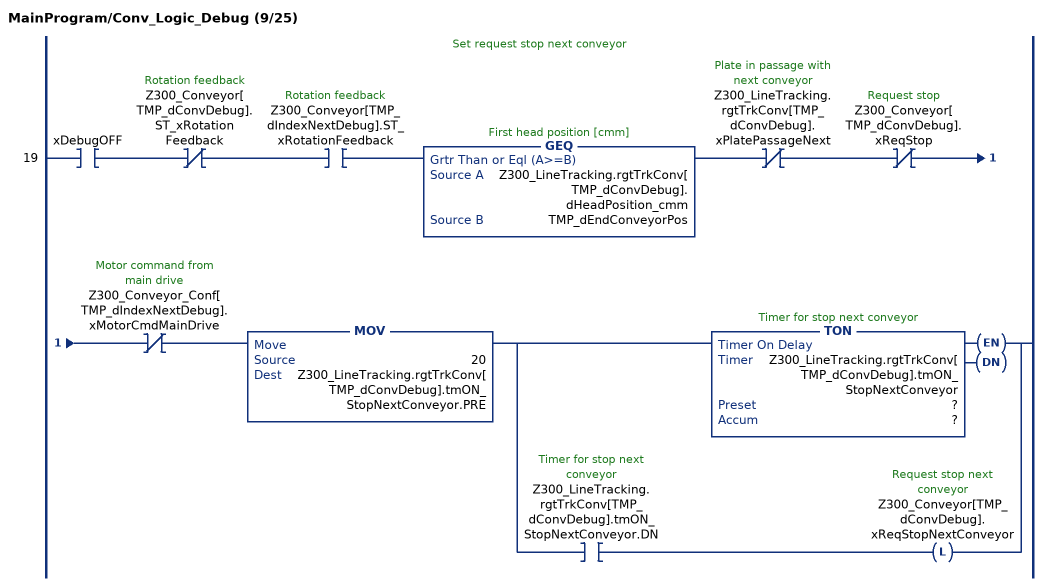
   // Set request stop next conveyor
   19: XIC(xDebugOFF)XIO(Z300_Conveyor[TMP_dConvDebug].ST_xRotationFeedback)XIC(Z300_Conveyor[TMP_dIndexNextDebug].ST_xRotationFeedback)GEQ(Z300_LineTracking.rgtTrkConv[TMP_dConvDebug].dHeadPosition_cmm,TMP_dEndConveyorPos)XIO(Z300_LineTracking.rgtTrkConv[TMP_dConvDebug].xPlatePassageNext)XIO(Z300_Conveyor[TMP_dConvDebug].xReqStop)XIO(Z300_Conveyor_Conf[TMP_dIndexNextDebug].xMotorCmdMainDrive)MOV(20,Z300_LineTracking.rgtTrkConv[TMP_dConvDebug].tmON_StopNextConveyor.PRE)[TON(Z300_LineTracking.rgtTrkConv[TMP_dConvDebug].tmON_StopNextConveyor,?,?) ,XIC(Z300_LineTracking.rgtTrkConv[TMP_dConvDebug].tmON_StopNextConveyor.DN) OTL(Z300_Conveyor[TMP_dConvDebug].xReqStopNextConveyor) ];
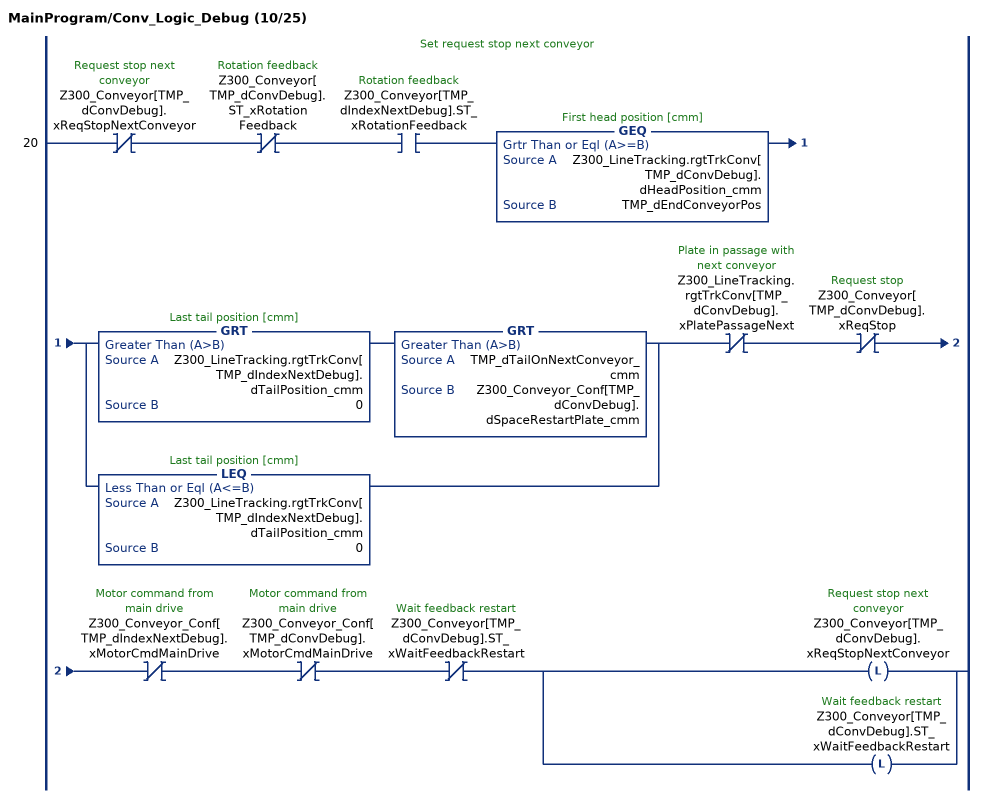
   // Set request stop next conveyor
   20: XIO(Z300_Conveyor[TMP_dConvDebug].xReqStopNextConveyor)XIO(Z300_Conveyor[TMP_dConvDebug].ST_xRotationFeedback)XIC(Z300_Conveyor[TMP_dIndexNextDebug].ST_xRotationFeedback)GEQ(Z300_LineTracking.rgtTrkConv[TMP_dConvDebug].dHeadPosition_cmm,TMP_dEndConveyorPos)[GRT(Z300_LineTracking.rgtTrkConv[TMP_dIndexNextDebug].dTailPosition_cmm,0) GRT(TMP_dTailOnNextConveyor_cmm,Z300_Conveyor_Conf[TMP_dConvDebug].dSpaceRestartPlate_cmm) ,LEQ(Z300_LineTracking.rgtTrkConv[TMP_dIndexNextDebug].dTailPosition_cmm,0) ]XIO(Z300_LineTracking.rgtTrkConv[TMP_dConvDebug].xPlatePassageNext)XIO(Z300_Conveyor[TMP_dConvDebug].xReqStop)XIO(Z300_Conveyor_Conf[TMP_dIndexNextDebug].xMotorCmdMainDrive)XIO(Z300_Conveyor_Conf[TMP_dConvDebug].xMotorCmdMainDrive)XIO(Z300_Conveyor[TMP_dConvDebug].ST_xWaitFeedbackRestart)[OTL(Z300_Conveyor[TMP_dConvDebug].xReqStopNextConveyor) ,OTL(Z300_Conveyor[TMP_dConvDebug].ST_xWaitFeedbackRestart) ];
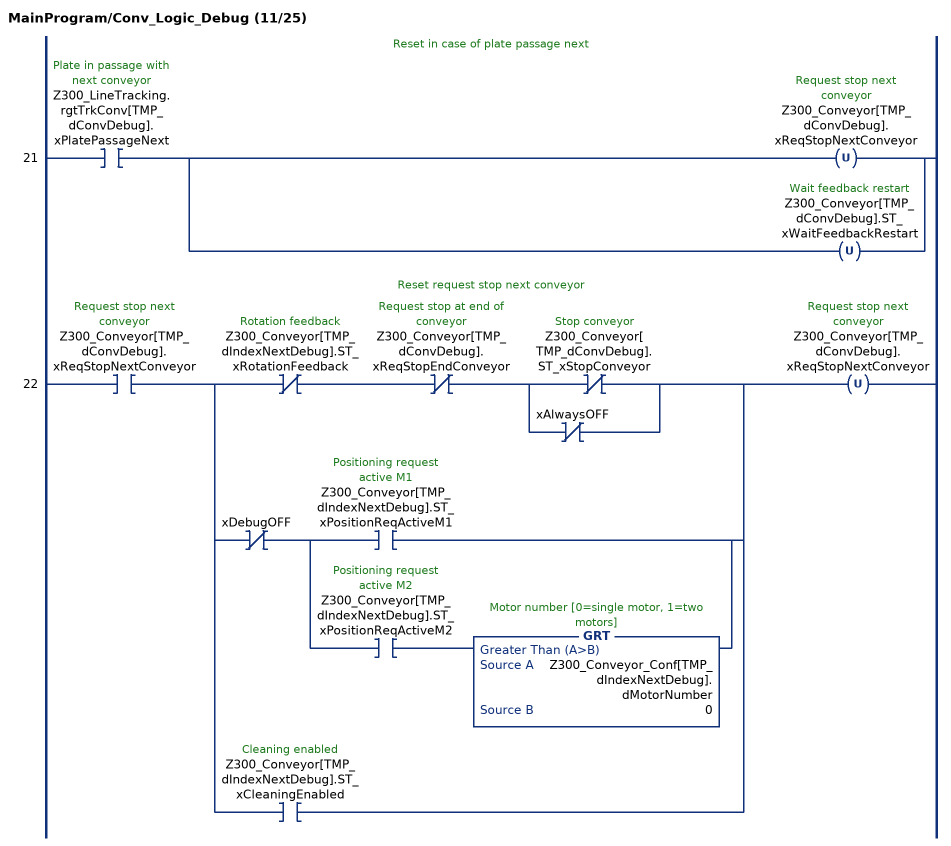
   // Reset in case of plate passage next
   21: XIC(Z300_LineTracking.rgtTrkConv[TMP_dConvDebug].xPlatePassageNext)[OTU(Z300_Conveyor[TMP_dConvDebug].xReqStopNextConveyor) ,OTU(Z300_Conveyor[TMP_dConvDebug].ST_xWaitFeedbackRestart) ];
   // Reset request stop next conveyor
   22: XIC(Z300_Conveyor[TMP_dConvDebug].xReqStopNextConveyor)[XIO(Z300_Conveyor[TMP_dIndexNextDebug].ST_xRotationFeedback) XIO(Z300_Conveyor[TMP_dConvDebug].xReqStopEndConveyor) [XIO(Z300_Conveyor[TMP_dConvDebug].ST_xStopConveyor) ,XIO(xAlwaysOFF) ] ,XIO(xDebugOFF) [XIC(Z300_Conveyor[TMP_dIndexNextDebug].ST_xPositionReqActiveM1) ,XIC(Z300_Conveyor[TMP_dIndexNextDebug].ST_xPositionReqActiveM2) GRT(Z300_Conveyor_Conf[TMP_dIndexNextDebug].dMotorNumber,0) ] ,XIC(Z300_Conveyor[TMP_dIndexNextDebug].ST_xCleaningEnabled) ]OTU(Z300_Conveyor[TMP_dConvDebug].xReqStopNextConveyor);
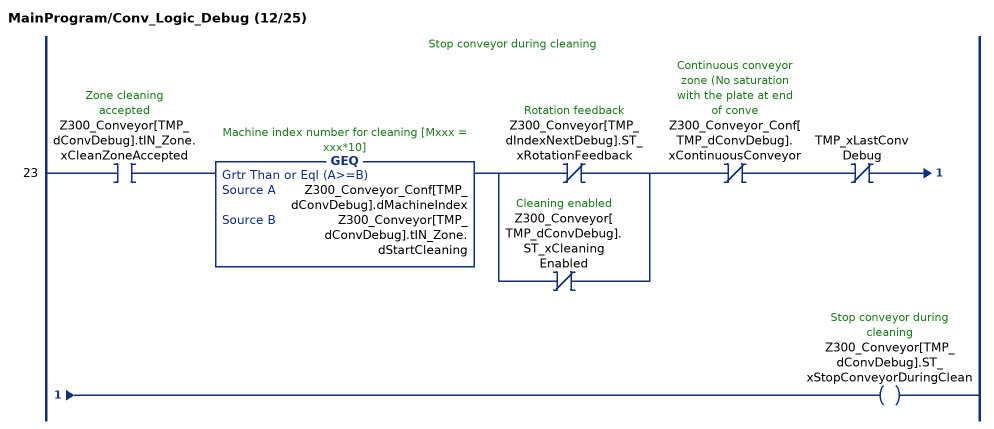
   // Stop conveyor during cleaning
   23: XIC(Z300_Conveyor[TMP_dConvDebug].tIN_Zone.xCleanZoneAccepted)GEQ(Z300_Conveyor_Conf[TMP_dConvDebug].dMachineIndex,Z300_Conveyor[TMP_dConvDebug].tIN_Zone.dStartCleaning)[XIO(Z300_Conveyor[TMP_dIndexNextDebug].ST_xRotationFeedback) ,XIO(Z300_Conveyor[TMP_dConvDebug].ST_xCleaningEnabled) ]XIO(Z300_Conveyor_Conf[TMP_dConvDebug].xContinuousConveyor)XIO(TMP_xLastConvDebug)OTE(Z300_Conveyor[TMP_dConvDebug].ST_xStopConveyorDuringClean);
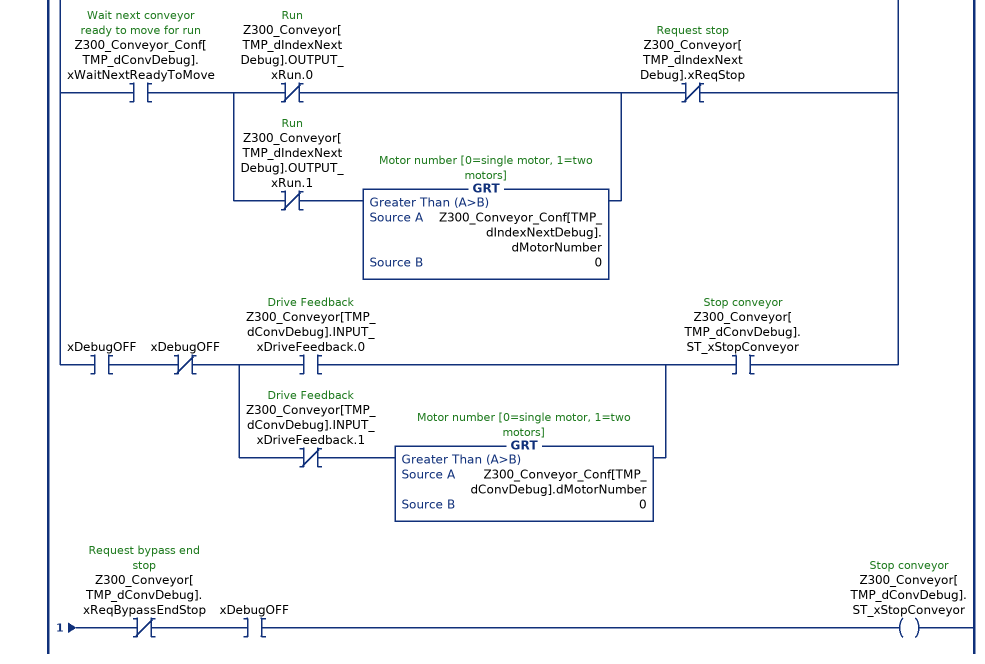
   // Stop conveyor
   24: [[XIC(Z300_LineTracking.rgtTrkConv[TMP_dConvDebug].xPlatePassagePrevious) [XIO(Z300_Conveyor[TMP_dIndexPreviousDebug].ST_xOutputEnable) ,XIC(Z300_Conveyor[TMP_dIndexPreviousDebug].ST_xWaitStopConveyor) ,XIC(xAlwaysOFF) XIC(Z300_Conveyor[TMP_dIndexPreviousDebug].xReqStop) ] ,XIC(Z300_LineTracking.rgtTrkConv[TMP_dConvDebug].xPlatePassageNext) XIO(TMP_xLastConvDebug) [XIO(Z300_Conveyor[TMP_dIndexNextDebug].ST_xOutMotorRun) ,XIO(Z300_Conveyor[TMP_dIndexNextDebug].INPUT_xSafetyConveyor) ] ,XIC(Z300_Conveyor[TMP_dConvDebug].ST_xStopPlateAtEndConveyor) ,XIC(Z300_Conveyor[TMP_dConvDebug].xReqStopNextConveyor) XIC(Z300_Conveyor[TMP_dIndexNextDebug].ST_xRotationFeedback) ,XIC(Z300_Conveyor[TMP_dConvDebug].ST_xStopConveyorDuringClean) ] [XIO(Z300_Conveyor_Conf[TMP_dConvDebug].xContinuousConveyor) ,XIC(Z300_Conveyor_Conf[TMP_dConvDebug].xEnableStopPlateContinuousZone) XIC(Z300_Conveyor[TMP_dConvDebug].xReqStopEndConveyor) ] ,XIC(Z300_Conveyor[TMP_dIndexPreviousDebug].xReqStopNextConveyor) XIO(Z300_Conveyor[TMP_dConvDebug].tIN_Zone.xCleanZoneAccepted) XIO(Z300_LineTracking.rgtTrkConv[TMP_dConvDebug].xGlassPresence) ,XIC(Z300_Conveyor_Conf[TMP_dConvDebug].xWaitNextReadyToMove) [XIO(Z300_Conveyor[TMP_dIndexNextDebug].OUTPUT_xRun.0) ,XIO(Z300_Conveyor[TMP_dIndexNextDebug].OUTPUT_xRun.1) GRT(Z300_Conveyor_Conf[TMP_dIndexNextDebug].dMotorNumber,0) ] XIO(Z300_Conveyor[TMP_dIndexNextDebug].xReqStop) ,XIC(xDebugOFF) XIO(xDebugOFF) [XIC(Z300_Conveyor[TMP_dConvDebug].INPUT_xDriveFeedback.0) ,XIO(Z300_Conveyor[TMP_dConvDebug].INPUT_xDriveFeedback.1) GRT(Z300_Conveyor_Conf[TMP_dConvDebug].dMotorNumber,0) ] XIC(Z300_Conveyor[TMP_dConvDebug].ST_xStopConveyor) ]XIO(Z300_Conveyor[TMP_dConvDebug].xReqBypassEndStop)XIC(xDebugOFF)OTE(Z300_Conveyor[TMP_dConvDebug].ST_xStopConveyor);
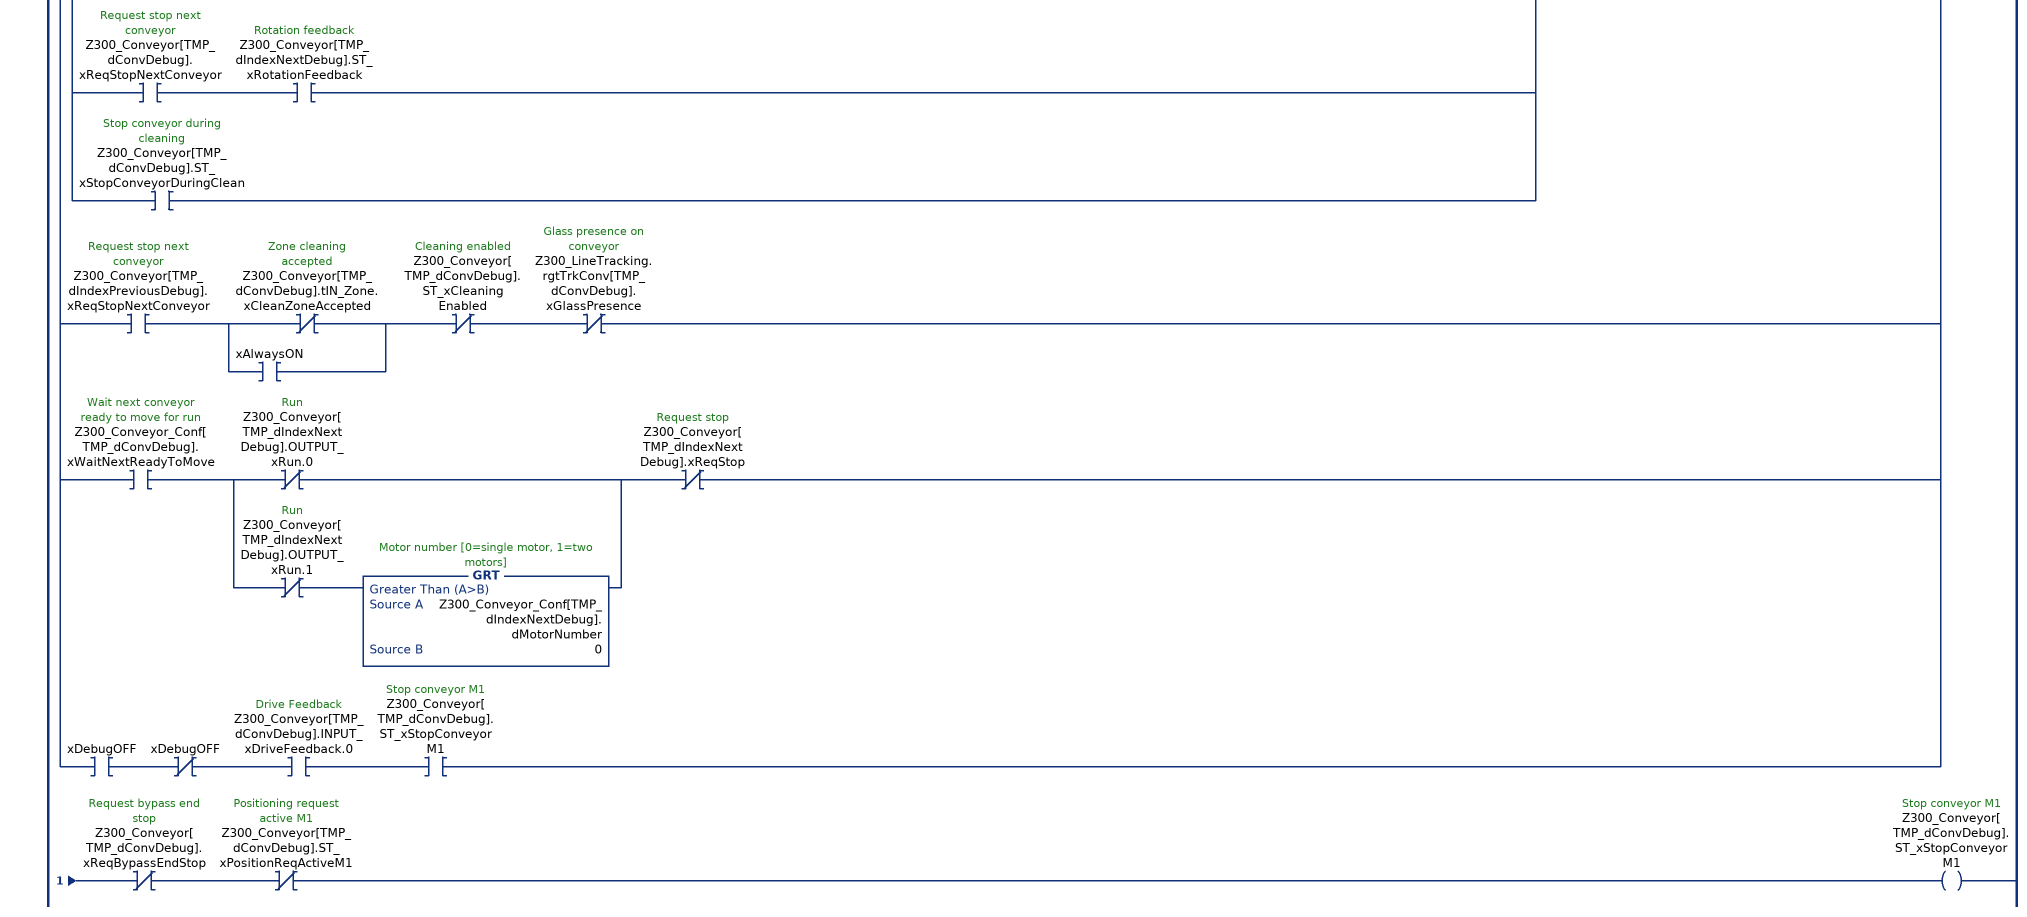
   // Stop conveyor M1
   // Monterrey VF2 - If this is conveyor after drop section I stop convveyor just if tail is under certain quote
   25: [[XIC(Z300_LineTracking.rgtTrkConv[TMP_dConvDebug].xPlatePassagePrevious) [XIO(Z300_Conveyor[TMP_dIndexPreviousDebug].ST_xOutputEnable) ,XIC(xDebugOFF) XIO(Z300_Conveyor[TMP_dIndexPreviousDebug].tmON_DelayReadyToMove[0].DN) ,XIC(Z300_Conveyor[TMP_dIndexPreviousDebug].ST_xInitialCondition) ,XIC(xDebugOFF) XIC(Z300_Conveyor[TMP_dIndexPreviousDebug].ST_xWaitStopConveyor) ,XIC(xAlwaysOFF) XIC(Z300_Conveyor[TMP_dIndexPreviousDebug].xReqStop) ] ,XIC(Z300_LineTracking.rgtTrkConv[TMP_dConvDebug].xPlatePassageNext) XIO(TMP_xLastConvDebug) [XIO(xDebugOFF) [EQU(TMP_dConvDebug,12) LES(Z300_LineTracking.rgtTrkConv[TMP_dConvDebug].dTailPosition_cmm,4100000) ,NEQ(TMP_dConvDebug,12) ] XIO(xDebugOFF) [XIO(Z300_Conveyor[TMP_dIndexNextDebug].ST_xOutMotorRun) ,XIC(xAlwaysON) ] XIO(Z300_Conveyor[TMP_dIndexNextDebug].ST_rgxConveyorOutRunSgm.0) XIO(Z300_Conveyor[TMP_dIndexNextDebug].ST_rgxConveyorOutRunSgm.1) ,XIO(Z300_Conveyor[TMP_dIndexNextDebug].INPUT_xSafetyConveyor) ] ,XIC(Z300_Conveyor[TMP_dConvDebug].ST_xStopPlateAtEndConveyor) XIO(Z300_Conveyor[TMP_dConvDebug].xReqBypassEndConveyorM1) ,XIC(Z300_Conveyor[TMP_dConvDebug].xReqStopNextConveyor) XIC(Z300_Conveyor[TMP_dIndexNextDebug].ST_xRotationFeedback) ,XIC(Z300_Conveyor[TMP_dConvDebug].ST_xStopConveyorDuringClean) ] [XIO(Z300_Conveyor_Conf[TMP_dConvDebug].xContinuousConveyor) ,XIC(Z300_Conveyor_Conf[TMP_dConvDebug].xEnableStopPlateContinuousZone) XIC(Z300_Conveyor[TMP_dConvDebug].xReqStopEndConveyor) ] ,XIC(Z300_Conveyor[TMP_dIndexPreviousDebug].xReqStopNextConveyor) [XIO(Z300_Conveyor[TMP_dConvDebug].tIN_Zone.xCleanZoneAccepted) ,XIC(xAlwaysON) ] XIO(Z300_Conveyor[TMP_dConvDebug].ST_xCleaningEnabled) XIO(Z300_LineTracking.rgtTrkConv[TMP_dConvDebug].xGlassPresence) ,XIC(Z300_Conveyor_Conf[TMP_dConvDebug].xWaitNextReadyToMove) [XIO(Z300_Conveyor[TMP_dIndexNextDebug].OUTPUT_xRun.0) ,XIO(Z300_Conveyor[TMP_dIndexNextDebug].OUTPUT_xRun.1) GRT(Z300_Conveyor_Conf[TMP_dIndexNextDebug].dMotorNumber,0) ] XIO(Z300_Conveyor[TMP_dIndexNextDebug].xReqStop) ,XIC(xDebugOFF) XIO(xDebugOFF) XIC(Z300_Conveyor[TMP_dConvDebug].INPUT_xDriveFeedback.0) XIC(Z300_Conveyor[TMP_dConvDebug].ST_xStopConveyorM1) ]XIO(Z300_Conveyor[TMP_dConvDebug].xReqBypassEndStop)XIO(Z300_Conveyor[TMP_dConvDebug].ST_xPositionReqActiveM1)OTE(Z300_Conveyor[TMP_dConvDebug].ST_xStopConveyorM1);
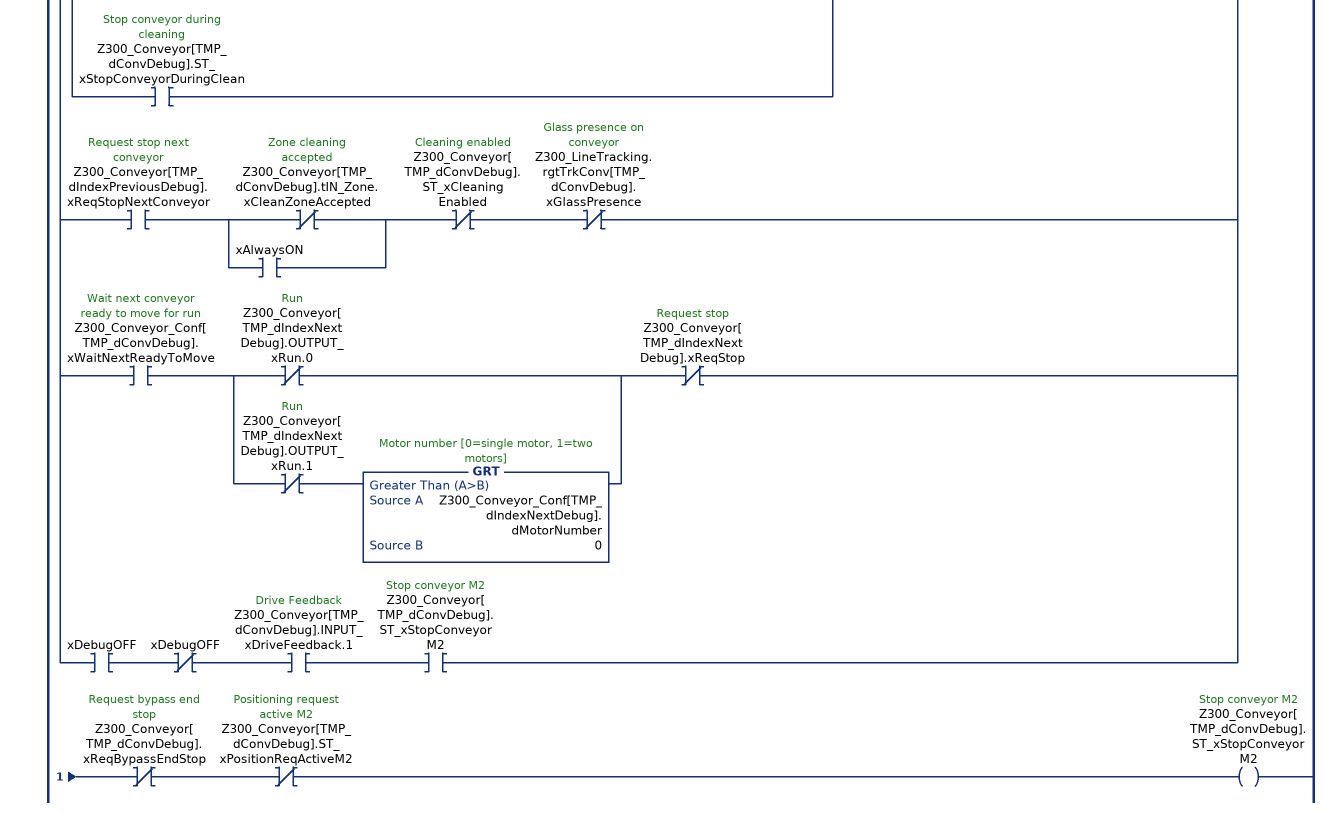
   // Stop conveyor M2
   // Monterrey VF2 - If this is conveyor after drop section I stop convveyor just if tail is under certain quote
   26: [[XIC(Z300_LineTracking.rgtTrkConv[TMP_dConvDebug].xPlatePassagePrevious) [XIO(Z300_Conveyor[TMP_dIndexPreviousDebug].ST_xOutputEnable) ,XIC(xDebugOFF) XIO(Z300_Conveyor[TMP_dIndexPreviousDebug].tmON_DelayReadyToMove[1].DN) ,XIC(Z300_Conveyor[TMP_dIndexPreviousDebug].ST_xInitialCondition) ,XIC(xDebugOFF) XIC(Z300_Conveyor[TMP_dIndexPreviousDebug].ST_xWaitStopConveyor) ,XIC(xAlwaysOFF) XIC(Z300_Conveyor[TMP_dIndexPreviousDebug].xReqStop) ] ,XIC(Z300_LineTracking.rgtTrkConv[TMP_dConvDebug].xPlatePassageNext) XIO(TMP_xLastConvDebug) [[XIO(Z300_Conveyor[TMP_dIndexNextDebug].ST_xOutMotorRun) ,XIC(xAlwaysON) ] XIO(Z300_Conveyor[TMP_dIndexNextDebug].ST_rgxConveyorOutRunSgm.0) XIO(Z300_Conveyor[TMP_dIndexNextDebug].ST_rgxConveyorOutRunSgm.1) ,XIO(Z300_Conveyor[TMP_dIndexNextDebug].INPUT_xSafetyConveyor) ] ,XIC(Z300_Conveyor[TMP_dConvDebug].ST_xStopPlateAtEndConveyor) XIO(Z300_Conveyor[TMP_dConvDebug].xReqBypassEndConveyorM2) ,XIC(Z300_Conveyor[TMP_dConvDebug].xReqStopNextConveyor) XIC(Z300_Conveyor[TMP_dIndexNextDebug].ST_xRotationFeedback) ,XIC(Z300_Conveyor[TMP_dConvDebug].ST_xStopConveyorDuringClean) ] [XIO(Z300_Conveyor_Conf[TMP_dConvDebug].xContinuousConveyor) ,XIC(Z300_Conveyor_Conf[TMP_dConvDebug].xEnableStopPlateContinuousZone) XIC(Z300_Conveyor[TMP_dConvDebug].xReqStopEndConveyor) ] ,XIC(Z300_Conveyor[TMP_dIndexPreviousDebug].xReqStopNextConveyor) [XIO(Z300_Conveyor[TMP_dConvDebug].tIN_Zone.xCleanZoneAccepted) ,XIC(xAlwaysON) ] XIO(Z300_Conveyor[TMP_dConvDebug].ST_xCleaningEnabled) XIO(Z300_LineTracking.rgtTrkConv[TMP_dConvDebug].xGlassPresence) ,XIC(Z300_Conveyor_Conf[TMP_dConvDebug].xWaitNextReadyToMove) [XIO(Z300_Conveyor[TMP_dIndexNextDebug].OUTPUT_xRun.0) ,XIO(Z300_Conveyor[TMP_dIndexNextDebug].OUTPUT_xRun.1) GRT(Z300_Conveyor_Conf[TMP_dIndexNextDebug].dMotorNumber,0) ] XIO(Z300_Conveyor[TMP_dIndexNextDebug].xReqStop) ,XIC(xDebugOFF) XIO(xDebugOFF) XIC(Z300_Conveyor[TMP_dConvDebug].INPUT_xDriveFeedback.1) XIC(Z300_Conveyor[TMP_dConvDebug].ST_xStopConveyorM2) ]XIO(Z300_Conveyor[TMP_dConvDebug].xReqBypassEndStop)XIO(Z300_Conveyor[TMP_dConvDebug].ST_xPositionReqActiveM2)OTE(Z300_Conveyor[TMP_dConvDebug].ST_xStopConveyorM2);
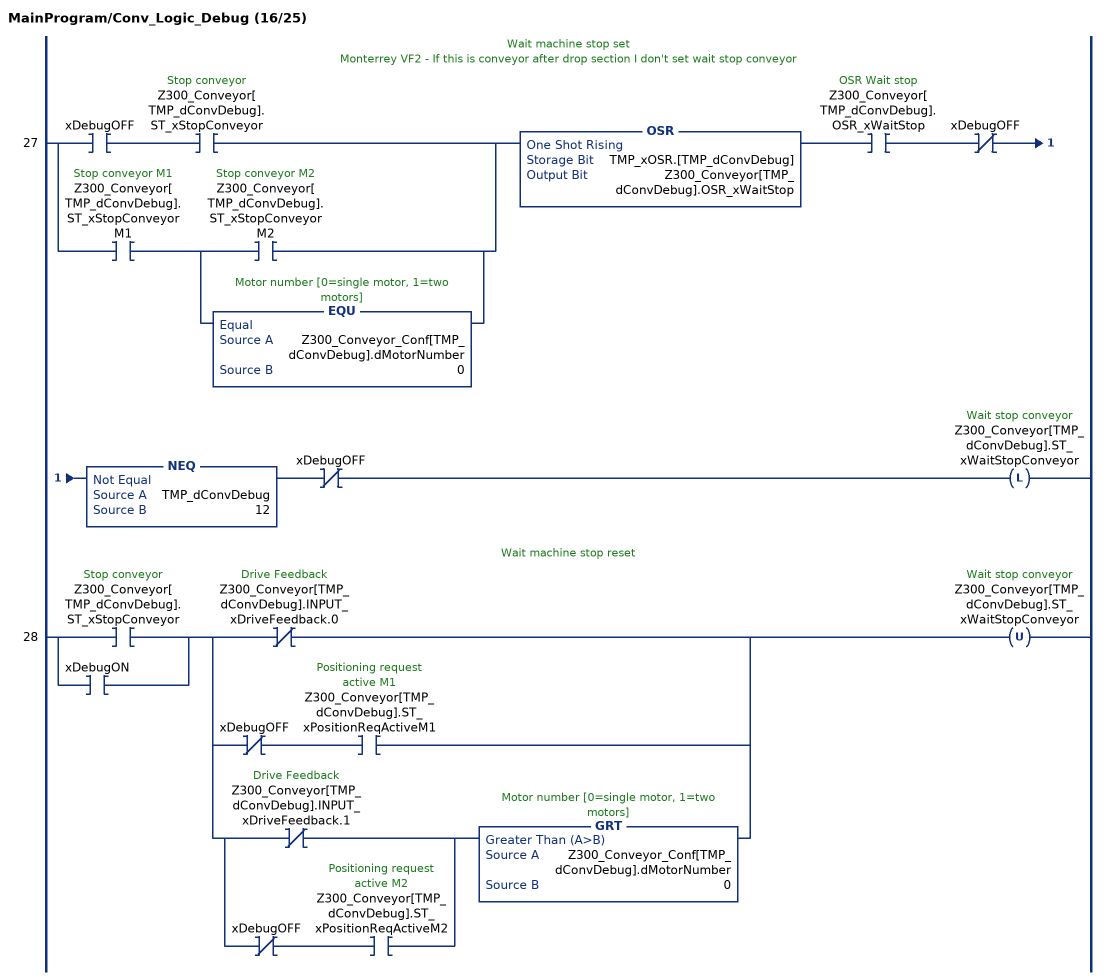
   // Wait machine stop set
   // Monterrey VF2 - If this is conveyor after drop section I don't set wait stop conveyor
   27: [XIC(xDebugOFF) XIC(Z300_Conveyor[TMP_dConvDebug].ST_xStopConveyor) ,XIC(Z300_Conveyor[TMP_dConvDebug].ST_xStopConveyorM1) [XIC(Z300_Conveyor[TMP_dConvDebug].ST_xStopConveyorM2) ,EQU(Z300_Conveyor_Conf[TMP_dConvDebug].dMotorNumber,0) ] ]OSR(TMP_xOSR.[TMP_dConvDebug],Z300_Conveyor[TMP_dConvDebug].OSR_xWaitStop)XIC(Z300_Conveyor[TMP_dConvDebug].OSR_xWaitStop)XIO(xDebugOFF)NEQ(TMP_dConvDebug,12)XIO(xDebugOFF)OTL(Z300_Conveyor[TMP_dConvDebug].ST_xWaitStopConveyor);
   // Wait machine stop reset
   28: [XIC(Z300_Conveyor[TMP_dConvDebug].ST_xStopConveyor) ,XIC(xDebugON) ][XIO(Z300_Conveyor[TMP_dConvDebug].INPUT_xDriveFeedback.0) ,XIO(xDebugOFF) XIC(Z300_Conveyor[TMP_dConvDebug].ST_xPositionReqActiveM1) ,[XIO(Z300_Conveyor[TMP_dConvDebug].INPUT_xDriveFeedback.1) ,XIO(xDebugOFF) XIC(Z300_Conveyor[TMP_dConvDebug].ST_xPositionReqActiveM2) ] GRT(Z300_Conveyor_Conf[TMP_dConvDebug].dMotorNumber,0) ]OTU(Z300_Conveyor[TMP_dConvDebug].ST_xWaitStopConveyor);
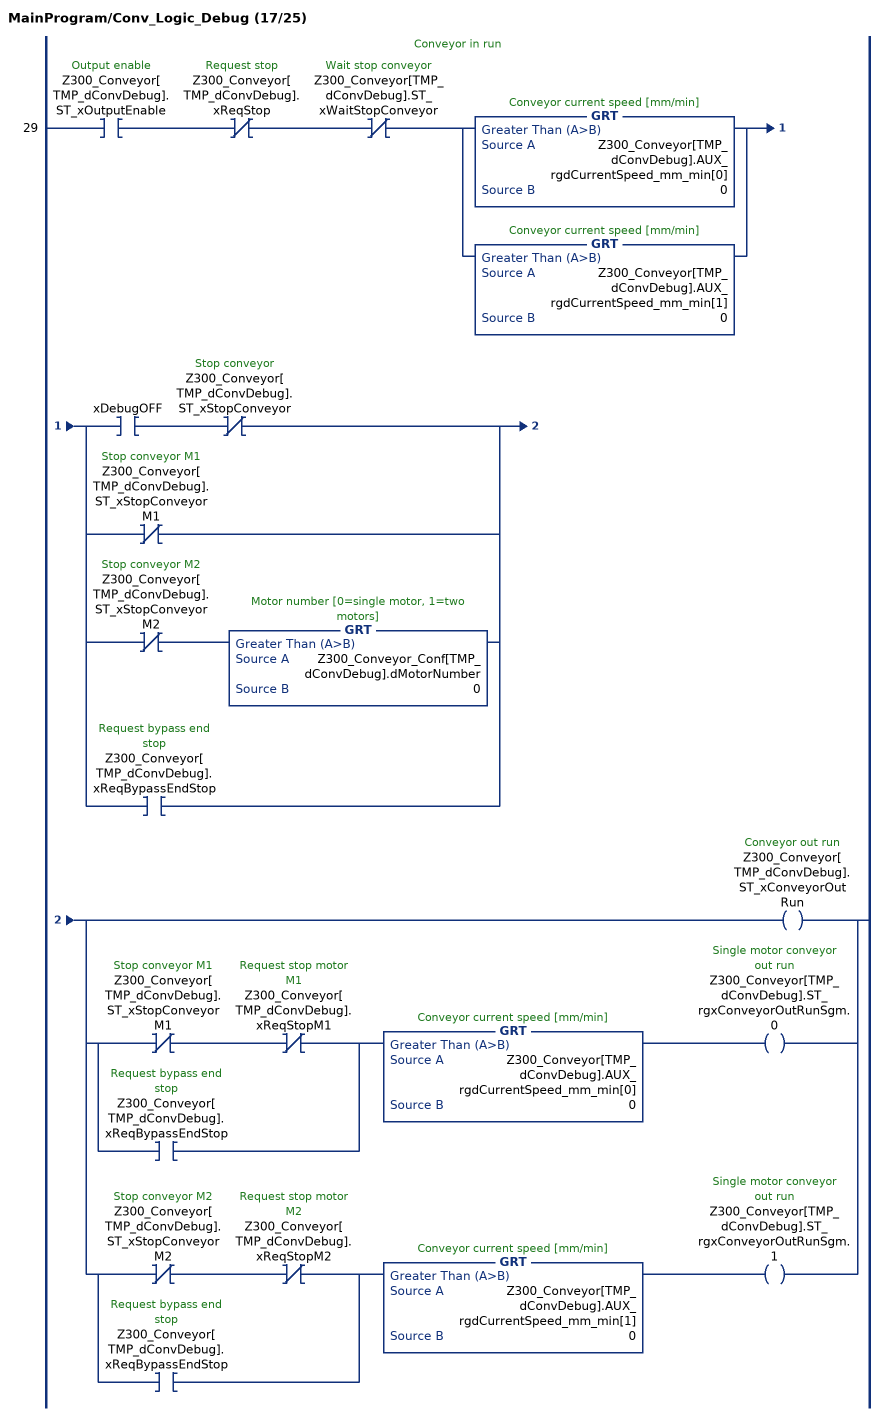
   // Conveyor in run
   29: XIC(Z300_Conveyor[TMP_dConvDebug].ST_xOutputEnable)XIO(Z300_Conveyor[TMP_dConvDebug].xReqStop)XIO(Z300_Conveyor[TMP_dConvDebug].ST_xWaitStopConveyor)[GRT(Z300_Conveyor[TMP_dConvDebug].AUX_rgdCurrentSpeed_mm_min[0],0) ,GRT(Z300_Conveyor[TMP_dConvDebug].AUX_rgdCurrentSpeed_mm_min[1],0) ][XIC(xDebugOFF) XIO(Z300_Conveyor[TMP_dConvDebug].ST_xStopConveyor) ,XIO(Z300_Conveyor[TMP_dConvDebug].ST_xStopConveyorM1) ,XIO(Z300_Conveyor[TMP_dConvDebug].ST_xStopConveyorM2) GRT(Z300_Conveyor_Conf[TMP_dConvDebug].dMotorNumber,0) ,XIC(Z300_Conveyor[TMP_dConvDebug].xReqBypassEndStop) ][OTE(Z300_Conveyor[TMP_dConvDebug].ST_xConveyorOutRun) ,[XIO(Z300_Conveyor[TMP_dConvDebug].ST_xStopConveyorM1) XIO(Z300_Conveyor[TMP_dConvDebug].xReqStopM1) ,XIC(Z300_Conveyor[TMP_dConvDebug].xReqBypassEndStop) ] GRT(Z300_Conveyor[TMP_dConvDebug].AUX_rgdCurrentSpeed_mm_min[0],0) OTE(Z300_Conveyor[TMP_dConvDebug].ST_rgxConveyorOutRunSgm.0) ,[XIO(Z300_Conveyor[TMP_dConvDebug].ST_xStopConveyorM2) XIO(Z300_Conveyor[TMP_dConvDebug].xReqStopM2) ,XIC(Z300_Conveyor[TMP_dConvDebug].xReqBypassEndStop) ] GRT(Z300_Conveyor[TMP_dConvDebug].AUX_rgdCurrentSpeed_mm_min[1],0) OTE(Z300_Conveyor[TMP_dConvDebug].ST_rgxConveyorOutRunSgm.1) ];
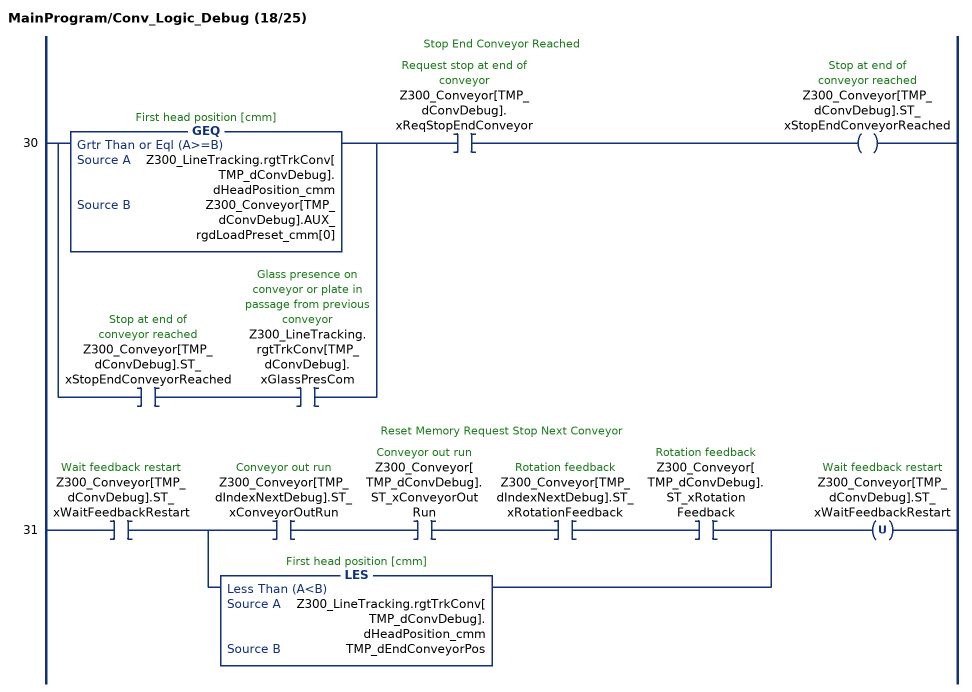
   // Stop End Conveyor Reached
   30: [GEQ(Z300_LineTracking.rgtTrkConv[TMP_dConvDebug].dHeadPosition_cmm,Z300_Conveyor[TMP_dConvDebug].AUX_rgdLoadPreset_cmm[0]) ,XIC(Z300_Conveyor[TMP_dConvDebug].ST_xStopEndConveyorReached) XIC(Z300_LineTracking.rgtTrkConv[TMP_dConvDebug].xGlassPresCom) ]XIC(Z300_Conveyor[TMP_dConvDebug].xReqStopEndConveyor)OTE(Z300_Conveyor[TMP_dConvDebug].ST_xStopEndConveyorReached);
   // Reset Memory Request Stop Next Conveyor
   31: XIC(Z300_Conveyor[TMP_dConvDebug].ST_xWaitFeedbackRestart)[XIC(Z300_Conveyor[TMP_dIndexNextDebug].ST_xConveyorOutRun) XIC(Z300_Conveyor[TMP_dConvDebug].ST_xConveyorOutRun) XIC(Z300_Conveyor[TMP_dIndexNextDebug].ST_xRotationFeedback) XIC(Z300_Conveyor[TMP_dConvDebug].ST_xRotationFeedback) ,LES(Z300_LineTracking.rgtTrkConv[TMP_dConvDebug].dHeadPosition_cmm,TMP_dEndConveyorPos) ]OTU(Z300_Conveyor[TMP_dConvDebug].ST_xWaitFeedbackRestart);
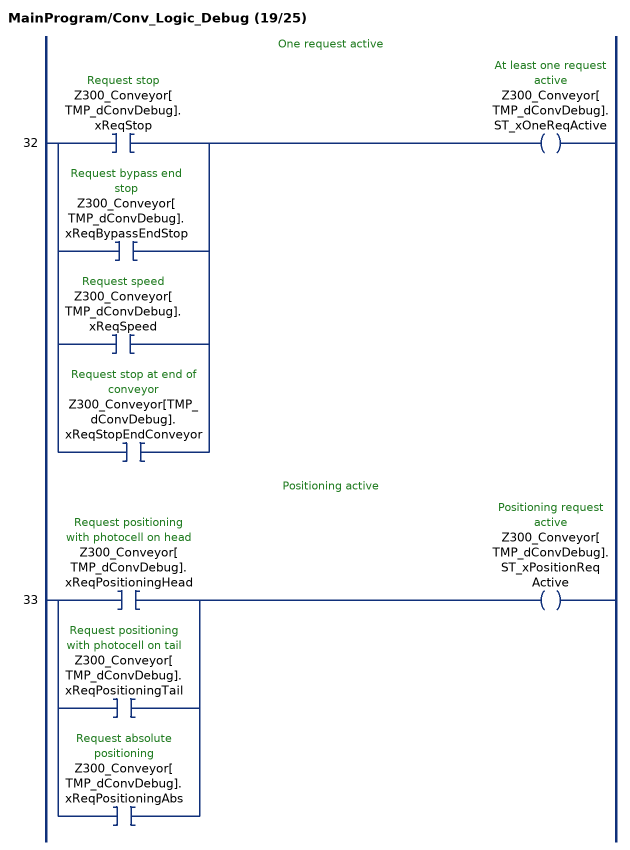
   // One request active
   32: [XIC(Z300_Conveyor[TMP_dConvDebug].xReqStop) ,XIC(Z300_Conveyor[TMP_dConvDebug].xReqBypassEndStop) ,XIC(Z300_Conveyor[TMP_dConvDebug].xReqSpeed) ,XIC(Z300_Conveyor[TMP_dConvDebug].xReqStopEndConveyor) ]OTE(Z300_Conveyor[TMP_dConvDebug].ST_xOneReqActive);
   // Positioning active
   33: [XIC(Z300_Conveyor[TMP_dConvDebug].xReqPositioningHead) ,XIC(Z300_Conveyor[TMP_dConvDebug].xReqPositioningTail) ,XIC(Z300_Conveyor[TMP_dConvDebug].xReqPositioningAbs) ]OTE(Z300_Conveyor[TMP_dConvDebug].ST_xPositionReqActive);
